// TIA Portal project "Delta_Praktika_P&P" (V17) (continued)
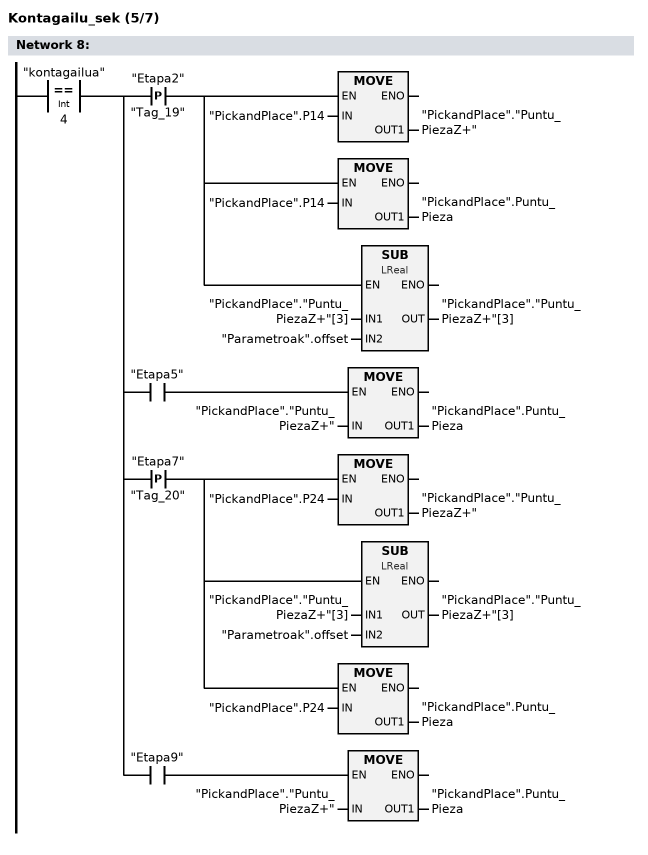
   RUNG wire#powerrail
      { S7_Templates := "SrcType := Int" } EQ_Contact(in1 := "kontagailua", in2 := 4)
      wire#w1
      P_Contact(operand := "Etapa2", bit := "Tag_19")
      wire#w2
      Move(in := "PickandPlace".P14, out1 => "PickandPlace"."Puntu_PiezaZ+")
   END_RUNG
   RUNG wire#w2
      Move(in := "PickandPlace".P14, out1 => "PickandPlace".Puntu_Pieza)
   END_RUNG
   RUNG wire#w2
      { S7_Templates := "SrcType := LReal" } Sub(in1 := "PickandPlace"."Puntu_PiezaZ+"[3], in2 := "Parametroak".offset, out => "PickandPlace"."Puntu_PiezaZ+"[3])
   END_RUNG
   RUNG wire#w1
      Contact( "Etapa5" )
      Move(in := "PickandPlace"."Puntu_PiezaZ+", out1 => "PickandPlace".Puntu_Pieza)
   END_RUNG
   RUNG wire#w1
      P_Contact(operand := "Etapa7", bit := "Tag_20")
      wire#w3
      Move(in := "PickandPlace".P24, out1 => "PickandPlace"."Puntu_PiezaZ+")
   END_RUNG
   RUNG wire#w3
      { S7_Templates := "SrcType := LReal" } Sub(in1 := "PickandPlace"."Puntu_PiezaZ+"[3], in2 := "Parametroak".offset, out => "PickandPlace"."Puntu_PiezaZ+"[3])
   END_RUNG
   RUNG wire#w3
      Move(in := "PickandPlace".P24, out1 => "PickandPlace".Puntu_Pieza)
   END_RUNG
   RUNG wire#w1
      Contact( "Etapa9" )
      Move(in := "PickandPlace"."Puntu_PiezaZ+", out1 => "PickandPlace".Puntu_Pieza)
   END_RUNG
   // the same network as SCL:
   #_w1 := "kontagailua" = 4;
   #_w2 := #_w1 AND "Etapa2" AND NOT "Tag_19";   // rising edge of "Etapa2"
   "Tag_19" := "Etapa2";
   IF #_w2 THEN
       "PickandPlace"."Puntu_PiezaZ+" := "PickandPlace".P14;
       "PickandPlace".Puntu_Pieza := "PickandPlace".P14;
       "PickandPlace"."Puntu_PiezaZ+"[3] := "PickandPlace"."Puntu_PiezaZ+"[3] - "Parametroak".offset;
   END_IF;
   IF #_w1 AND "Etapa5" THEN "PickandPlace".Puntu_Pieza := "PickandPlace"."Puntu_PiezaZ+"; END_IF;
   #_w3 := #_w1 AND "Etapa7" AND NOT "Tag_20";   // rising edge of "Etapa7"
   "Tag_20" := "Etapa7";
   IF #_w3 THEN
       "PickandPlace"."Puntu_PiezaZ+" := "PickandPlace".P24;
       "PickandPlace"."Puntu_PiezaZ+"[3] := "PickandPlace"."Puntu_PiezaZ+"[3] - "Parametroak".offset;
       "PickandPlace".Puntu_Pieza := "PickandPlace".P24;
   END_IF;
   IF #_w1 AND "Etapa9" THEN "PickandPlace".Puntu_Pieza := "PickandPlace"."Puntu_PiezaZ+"; END_IF;
END_REGION

REGION Network 9
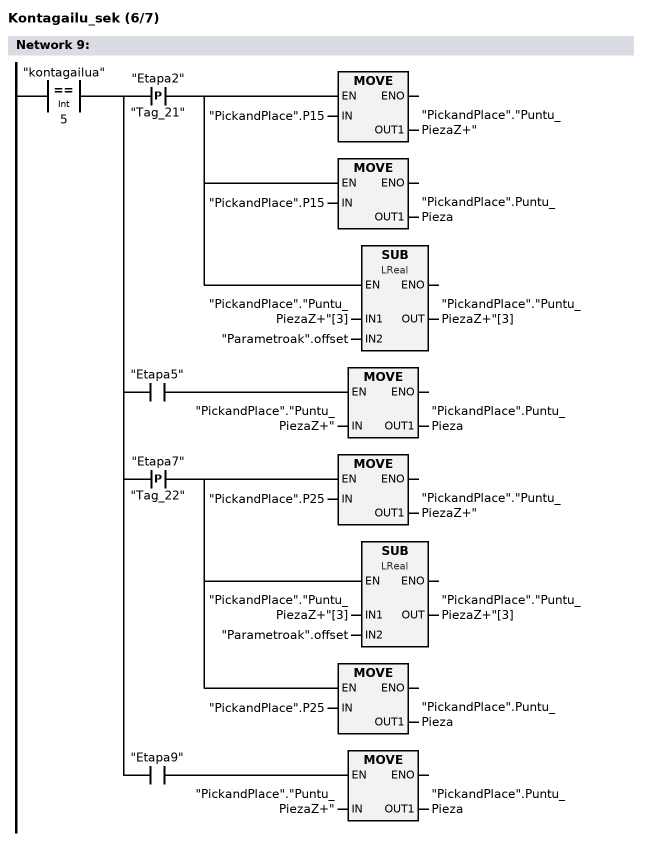
   RUNG wire#powerrail
      { S7_Templates := "SrcType := Int" } EQ_Contact(in1 := "kontagailua", in2 := 5)
      wire#w1
      P_Contact(operand := "Etapa2", bit := "Tag_21")
      wire#w2
      Move(in := "PickandPlace".P15, out1 => "PickandPlace"."Puntu_PiezaZ+")
   END_RUNG
   RUNG wire#w2
      Move(in := "PickandPlace".P15, out1 => "PickandPlace".Puntu_Pieza)
   END_RUNG
   RUNG wire#w2
      { S7_Templates := "SrcType := LReal" } Sub(in1 := "PickandPlace"."Puntu_PiezaZ+"[3], in2 := "Parametroak".offset, out => "PickandPlace"."Puntu_PiezaZ+"[3])
   END_RUNG
   RUNG wire#w1
      Contact( "Etapa5" )
      Move(in := "PickandPlace"."Puntu_PiezaZ+", out1 => "PickandPlace".Puntu_Pieza)
   END_RUNG
   RUNG wire#w1
      P_Contact(operand := "Etapa7", bit := "Tag_22")
      wire#w3
      Move(in := "PickandPlace".P25, out1 => "PickandPlace"."Puntu_PiezaZ+")
   END_RUNG
   RUNG wire#w3
      { S7_Templates := "SrcType := LReal" } Sub(in1 := "PickandPlace"."Puntu_PiezaZ+"[3], in2 := "Parametroak".offset, out => "PickandPlace"."Puntu_PiezaZ+"[3])
   END_RUNG
   RUNG wire#w3
      Move(in := "PickandPlace".P25, out1 => "PickandPlace".Puntu_Pieza)
   END_RUNG
   RUNG wire#w1
      Contact( "Etapa9" )
      Move(in := "PickandPlace"."Puntu_PiezaZ+", out1 => "PickandPlace".Puntu_Pieza)
   END_RUNG
   // the same network as SCL:
   #_w1 := "kontagailua" = 5;
   #_w2 := #_w1 AND "Etapa2" AND NOT "Tag_21";   // rising edge of "Etapa2"
   "Tag_21" := "Etapa2";
   IF #_w2 THEN
       "PickandPlace"."Puntu_PiezaZ+" := "PickandPlace".P15;
       "PickandPlace".Puntu_Pieza := "PickandPlace".P15;
       "PickandPlace"."Puntu_PiezaZ+"[3] := "PickandPlace"."Puntu_PiezaZ+"[3] - "Parametroak".offset;
   END_IF;
   IF #_w1 AND "Etapa5" THEN "PickandPlace".Puntu_Pieza := "PickandPlace"."Puntu_PiezaZ+"; END_IF;
   #_w3 := #_w1 AND "Etapa7" AND NOT "Tag_22";   // rising edge of "Etapa7"
   "Tag_22" := "Etapa7";
   IF #_w3 THEN
       "PickandPlace"."Puntu_PiezaZ+" := "PickandPlace".P25;
       "PickandPlace"."Puntu_PiezaZ+"[3] := "PickandPlace"."Puntu_PiezaZ+"[3] - "Parametroak".offset;
       "PickandPlace".Puntu_Pieza := "PickandPlace".P25;
   END_IF;
   IF #_w1 AND "Etapa9" THEN "PickandPlace".Puntu_Pieza := "PickandPlace"."Puntu_PiezaZ+"; END_IF;
END_REGION

REGION Network 10
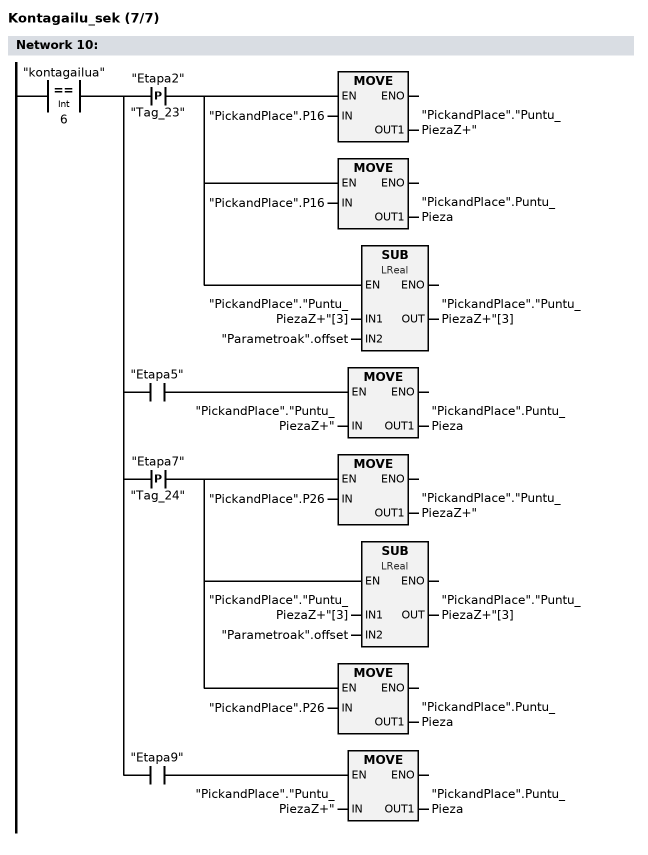
   RUNG wire#powerrail
      { S7_Templates := "SrcType := Int" } EQ_Contact(in1 := "kontagailua", in2 := 6)
      wire#w1
      P_Contact(operand := "Etapa2", bit := "Tag_23")
      wire#w2
      Move(in := "PickandPlace".P16, out1 => "PickandPlace"."Puntu_PiezaZ+")
   END_RUNG
   RUNG wire#w2
      Move(in := "PickandPlace".P16, out1 => "PickandPlace".Puntu_Pieza)
   END_RUNG
   RUNG wire#w2
      { S7_Templates := "SrcType := LReal" } Sub(in1 := "PickandPlace"."Puntu_PiezaZ+"[3], in2 := "Parametroak".offset, out => "PickandPlace"."Puntu_PiezaZ+"[3])
   END_RUNG
   RUNG wire#w1
      Contact( "Etapa5" )
      Move(in := "PickandPlace"."Puntu_PiezaZ+", out1 => "PickandPlace".Puntu_Pieza)
   END_RUNG
   RUNG wire#w1
      P_Contact(operand := "Etapa7", bit := "Tag_24")
      wire#w3
      Move(in := "PickandPlace".P26, out1 => "PickandPlace"."Puntu_PiezaZ+")
   END_RUNG
   RUNG wire#w3
      { S7_Templates := "SrcType := LReal" } Sub(in1 := "PickandPlace"."Puntu_PiezaZ+"[3], in2 := "Parametroak".offset, out => "PickandPlace"."Puntu_PiezaZ+"[3])
   END_RUNG
   RUNG wire#w3
      Move(in := "PickandPlace".P26, out1 => "PickandPlace".Puntu_Pieza)
   END_RUNG
   RUNG wire#w1
      Contact( "Etapa9" )
      Move(in := "PickandPlace"."Puntu_PiezaZ+", out1 => "PickandPlace".Puntu_Pieza)
   END_RUNG
   // the same network as SCL:
   #_w1 := "kontagailua" = 6;
   #_w2 := #_w1 AND "Etapa2" AND NOT "Tag_23";   // rising edge of "Etapa2"
   "Tag_23" := "Etapa2";
   IF #_w2 THEN
       "PickandPlace"."Puntu_PiezaZ+" := "PickandPlace".P16;
       "PickandPlace".Puntu_Pieza := "PickandPlace".P16;
       "PickandPlace"."Puntu_PiezaZ+"[3] := "PickandPlace"."Puntu_PiezaZ+"[3] - "Parametroak".offset;
   END_IF;
   IF #_w1 AND "Etapa5" THEN "PickandPlace".Puntu_Pieza := "PickandPlace"."Puntu_PiezaZ+"; END_IF;
   #_w3 := #_w1 AND "Etapa7" AND NOT "Tag_24";   // rising edge of "Etapa7"
   "Tag_24" := "Etapa7";
   IF #_w3 THEN
       "PickandPlace"."Puntu_PiezaZ+" := "PickandPlace".P26;
       "PickandPlace"."Puntu_PiezaZ+"[3] := "PickandPlace"."Puntu_PiezaZ+"[3] - "Parametroak".offset;
       "PickandPlace".Puntu_Pieza := "PickandPlace".P26;
   END_IF;
   IF #_w1 AND "Etapa9" THEN "PickandPlace".Puntu_Pieza := "PickandPlace"."Puntu_PiezaZ+"; END_IF;
END_REGION
END_FUNCTION

ORGANIZATION_BLOCK "Main"   // OB1, LAD, ProgramCycle
TITLE = "Main Program Sweep (Cycle)"
{ S7_Optimized_Access := 'TRUE' }
VERSION : 0.1
   VAR_INPUT
      Initial_Call : Bool;   // Initial call of this OB
      Remanence : Bool;   // =True, if remanent data are available
   END_VAR
BEGIN

REGION Network 1
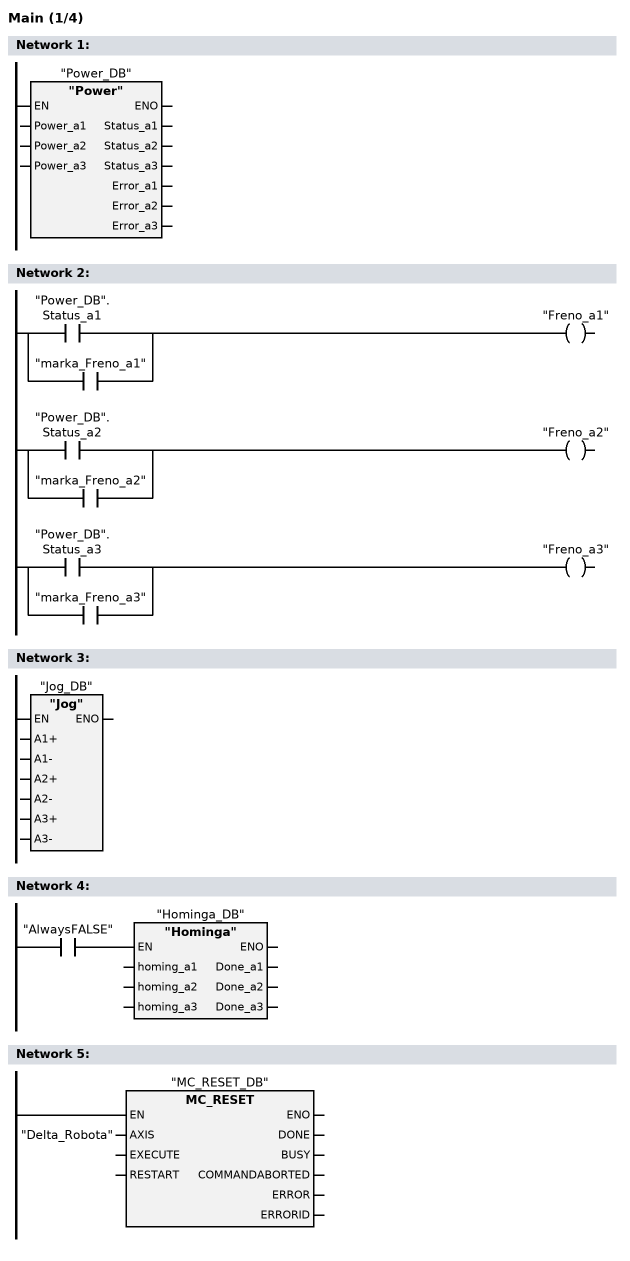
   RUNG wire#powerrail
      "Power_DB"(Power_a1 :=, Power_a2 :=, Power_a3 :=, Status_a1 =>, Status_a2 =>, Status_a3 =>, Error_a1 =>, Error_a2 =>, Error_a3 =>)
   END_RUNG
   // the same network as SCL:
   "Power_DB"();   // "Power"
END_REGION

REGION Network 2
   RUNG wire#powerrail
      Contact( "Power_DB".Status_a1 )
      wire#w1
      Coil( "Freno_a1" )
   END_RUNG
   RUNG wire#powerrail
      Contact( "marka_Freno_a1" )
   END_RUNG wire#w1
   RUNG wire#powerrail
      Contact( "Power_DB".Status_a2 )
      wire#w2
      Coil( "Freno_a2" )
   END_RUNG
   RUNG wire#powerrail
      Contact( "marka_Freno_a2" )
   END_RUNG wire#w2
   RUNG wire#powerrail
      Contact( "Power_DB".Status_a3 )
      wire#w3
      Coil( "Freno_a3" )
   END_RUNG
   RUNG wire#powerrail
      Contact( "marka_Freno_a3" )
   END_RUNG wire#w3
   // the same network as SCL:
   "Freno_a1" := "Power_DB".Status_a1 OR "marka_Freno_a1";
   "Freno_a2" := "Power_DB".Status_a2 OR "marka_Freno_a2";
   "Freno_a3" := "Power_DB".Status_a3 OR "marka_Freno_a3";
END_REGION

REGION Network 3
   RUNG wire#powerrail
      "Jog_DB"("A1+" :=, "A1-" :=, "A2+" :=, "A2-" :=, "A3+" :=, "A3-" :=)
   END_RUNG
   // the same network as SCL:
   "Jog_DB"();   // "Jog"
END_REGION

REGION Network 4
   RUNG wire#powerrail
      Contact( "AlwaysFALSE" )
      "Hominga_DB"(homing_a1 :=, homing_a2 :=, homing_a3 :=, Done_a1 =>, Done_a2 =>, Done_a3 =>)
   END_RUNG
   // the same network as SCL:
   IF "AlwaysFALSE" THEN
       "Hominga_DB"();   // "Hominga"
   END_IF;
END_REGION

REGION Network 5
   "MC_RESET_DB"(Axis := "Delta_Robota");   // MC_RESET
END_REGION

REGION Network 6
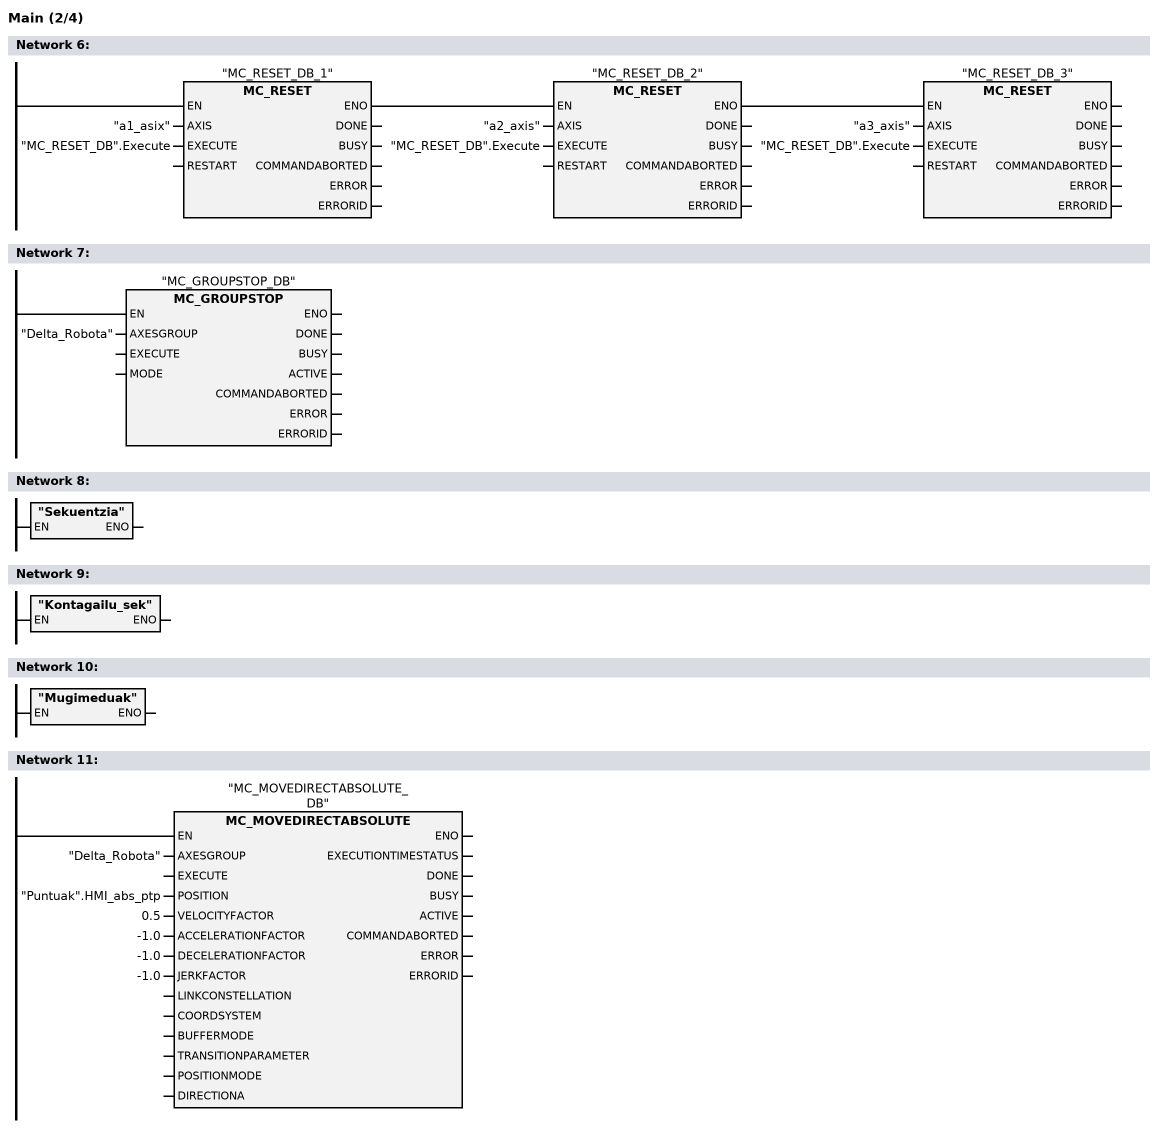
   // ENO of a box is taken as its EN; it also drops when the box reports an error
   "MC_RESET_DB_1"(Axis := "a1_asix", Execute := "MC_RESET_DB".Execute);   // MC_RESET
   "MC_RESET_DB_2"(Axis := "a2_axis", Execute := "MC_RESET_DB".Execute);   // MC_RESET
   "MC_RESET_DB_3"(Axis := "a3_axis", Execute := "MC_RESET_DB".Execute);   // MC_RESET
END_REGION

REGION Network 7
   "MC_GROUPSTOP_DB"(AxesGroup := "Delta_Robota");   // MC_GROUPSTOP
END_REGION

REGION Network 8
   RUNG wire#powerrail
      "Sekuentzia"()
   END_RUNG
   // the same network as SCL:
   "Sekuentzia"();
END_REGION

REGION Network 9
   RUNG wire#powerrail
      "Kontagailu_sek"()
   END_RUNG
   // the same network as SCL:
   "Kontagailu_sek"();
END_REGION

REGION Network 10
   RUNG wire#powerrail
      "Mugimeduak"()
   END_RUNG
   // the same network as SCL:
   "Mugimeduak"();
END_REGION

REGION Network 11
   "MC_MOVEDIRECTABSOLUTE_DB"(AxesGroup := "Delta_Robota",   // MC_MOVEDIRECTABSOLUTE
                           Position := "Puntuak".HMI_abs_ptp,
                           VelocityFactor := 0.5,
                           AccelerationFactor := -1.0,
                           DecelerationFactor := -1.0,
                           JerkFactor := -1.0);
END_REGION

REGION Network 12
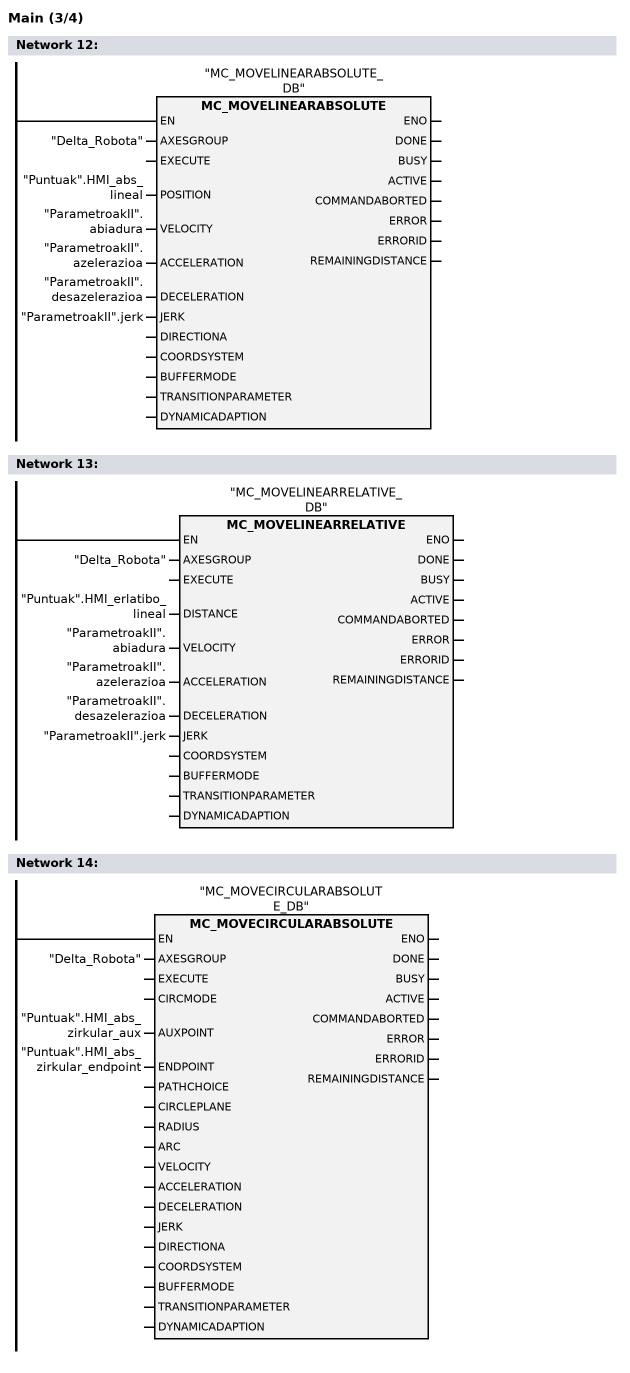
   "MC_MOVELINEARABSOLUTE_DB"(AxesGroup := "Delta_Robota",   // MC_MOVELINEARABSOLUTE
                           Position := "Puntuak".HMI_abs_lineal,
                           Velocity := "ParametroakII".abiadura,
                           Acceleration := "ParametroakII".azelerazioa,
                           Deceleration := "ParametroakII".desazelerazioa,
                           Jerk := "ParametroakII".jerk);
END_REGION

REGION Network 13
   "MC_MOVELINEARRELATIVE_DB"(AxesGroup := "Delta_Robota",   // MC_MOVELINEARRELATIVE
                           Distance := "Puntuak".HMI_erlatibo_lineal,
                           Velocity := "ParametroakII".abiadura,
                           Acceleration := "ParametroakII".azelerazioa,
                           Deceleration := "ParametroakII".desazelerazioa,
                           Jerk := "ParametroakII".jerk);
END_REGION

REGION Network 14
   "MC_MOVECIRCULARABSOLUTE_DB"(AxesGroup := "Delta_Robota",   // MC_MOVECIRCULARABSOLUTE
                           AuxPoint := "Puntuak".HMI_abs_zirkular_aux,
                           EndPoint := "Puntuak".HMI_abs_zirkular_endpoint);
END_REGION

REGION Network 15
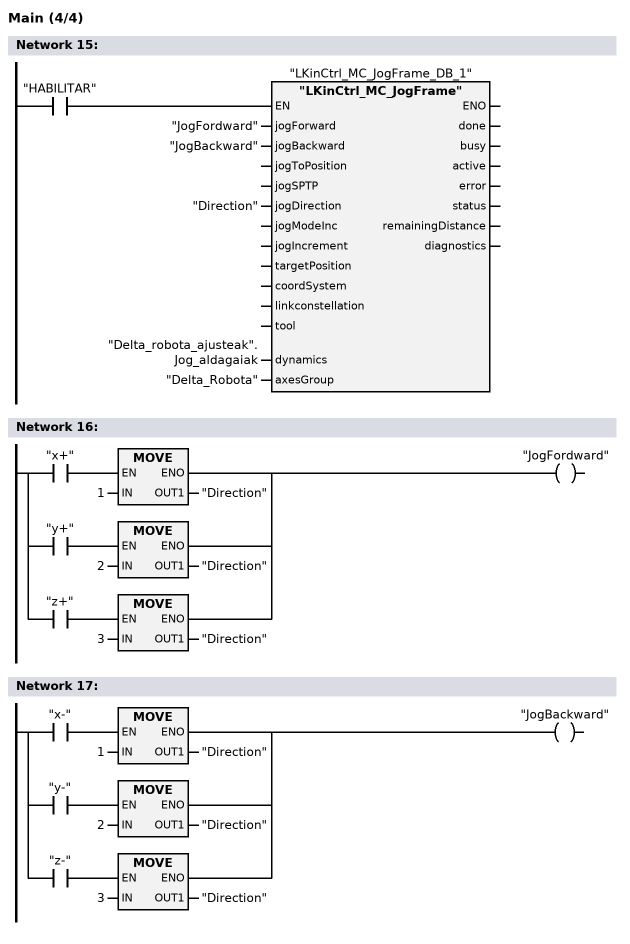
   RUNG wire#powerrail
      Contact( "HABILITAR" )
      "LKinCtrl_MC_JogFrame_DB_1"(jogForward := "JogFordward", jogBackward := "JogBackward", jogToPosition :=, jogSPTP :=, jogDirection := "Direction", jogModeInc :=, jogIncrement :=, targetPosition :=, coordSystem :=, linkconstellation :=, tool :=, dynamics := "Delta_robota_ajusteak".Jog_aldagaiak, axesGroup := "Delta_Robota", done =>, busy =>, active =>, error =>, status =>, remainingDistance =>, diagnostics =>)
   END_RUNG
   // the same network as SCL:
   IF "HABILITAR" THEN
       "LKinCtrl_MC_JogFrame_DB_1"(jogForward := "JogFordward",   // "LKinCtrl_MC_JogFrame"
                               jogBackward := "JogBackward",
                               jogDirection := "Direction",
                               dynamics := "Delta_robota_ajusteak".Jog_aldagaiak,
                               axesGroup := "Delta_Robota");
   END_IF;
END_REGION

REGION Network 16
   RUNG wire#powerrail
      Contact( "x+" )
      Move(in := 1, out1 => "Direction")
      wire#w1
      Coil( "JogFordward" )
   END_RUNG
   RUNG wire#powerrail
      Contact( "y+" )
      Move(in := 2, out1 => "Direction")
   END_RUNG wire#w1
   RUNG wire#powerrail
      Contact( "z+" )
      Move(in := 3, out1 => "Direction")
   END_RUNG wire#w1
   // the same network as SCL:
   IF "x+" THEN "Direction" := 1; END_IF;
   IF "y+" THEN "Direction" := 2; END_IF;
   IF "z+" THEN "Direction" := 3; END_IF;
   "JogFordward" := "x+" OR "y+" OR "z+";
END_REGION

REGION Network 17
   RUNG wire#powerrail
      Contact( "x-" )
      Move(in := 1, out1 => "Direction")
      wire#w1
      Coil( "JogBackward" )
   END_RUNG
   RUNG wire#powerrail
      Contact( "y-" )
      Move(in := 2, out1 => "Direction")
   END_RUNG wire#w1
   RUNG wire#powerrail
      Contact( "z-" )
      Move(in := 3, out1 => "Direction")
   END_RUNG wire#w1
   // the same network as SCL:
   IF "x-" THEN "Direction" := 1; END_IF;
   IF "y-" THEN "Direction" := 2; END_IF;
   IF "z-" THEN "Direction" := 3; END_IF;
   "JogBackward" := "x-" OR "y-" OR "z-";
END_REGION
END_ORGANIZATION_BLOCK

ORGANIZATION_BLOCK "Startup"   // OB100, LAD, Startup
TITLE = "Complete Restart"
{ S7_Optimized_Access := 'TRUE' }
VERSION : 0.1
   VAR_INPUT
      LostRetentive : Bool;   // True if retentive data are lost
      LostRTC : Bool;   // True if date and time are lost
   END_VAR
BEGIN

REGION Network 1
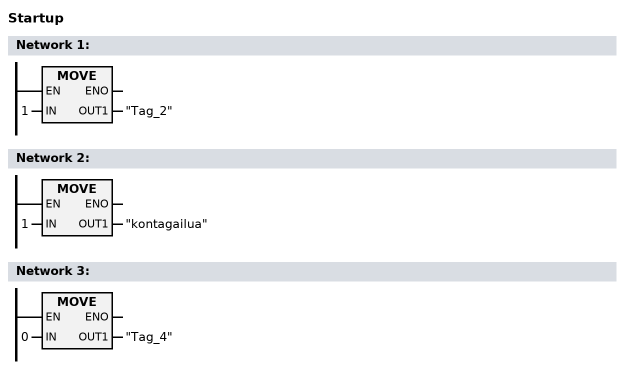
   RUNG wire#powerrail
      Move(in := 1, out1 => "Tag_2")
   END_RUNG
   // the same network as SCL:
   "Tag_2" := 1;
END_REGION

REGION Network 2
   RUNG wire#powerrail
      Move(in := 1, out1 => "kontagailua")
   END_RUNG
   // the same network as SCL:
   "kontagailua" := 1;
END_REGION

REGION Network 3
   RUNG wire#powerrail
      Move(in := 0, out1 => "Tag_4")
   END_RUNG
   // the same network as SCL:
   "Tag_4" := 0;
END_REGION
END_ORGANIZATION_BLOCK

(* ===== HMI "HMI_RT_1" =====
system functions are stored by id; their names below are inferred from use
connection "HMI_Conexión_2": ETHERNET, SMART_S7_1500_OMS

HMI tags "Tabla de variables estándar"
   "Delta_Robota_TcpInWcs_x_Position" : LReal = PLC Delta_Robota.TcpInWcs.x.Position, 1 s
   "Power_DB_Power_a1" : Bool = PLC Power_DB.Power_a1, 1 s
   "Jog_DB_A1+" : Bool = PLC Jog_DB.A1+, 1 s
   "a1_asix_ActualPosition" : LReal = PLC a1_asix.ActualPosition, 1 s
   "Power_DB_Power_a2" : Bool = PLC Power_DB.Power_a2, 1 s
   "Power_DB_Power_a3" : Bool = PLC Power_DB.Power_a3, 1 s
   "Tag_2" : Bool = PLC marka_Freno_a1 AT %M30.1, 1 s
   "Tag_3" : Bool = PLC marka_Freno_a2 AT %M30.2, 1 s
   "Tag_6" : Bool = PLC marka_Freno_a3 AT %M30.0, 1 s
   "Jog_DB_A1-" : Bool = PLC Jog_DB.A1-, 1 s
   "Jog_DB_A2+" : Bool = PLC Jog_DB.A2+, 1 s
   "Jog_DB_A2-" : Bool = PLC Jog_DB.A2-, 1 s
   "Jog_DB_A3+" : Bool = PLC Jog_DB.A3+, 1 s
   "Jog_DB_A3-" : Bool = PLC Jog_DB.A3-, 1 s
   "Tag_1" : Bool = PLC Freno_a1 AT %Q30.1, 1 s
   "Tag_4" : Bool = PLC Freno_a2 AT %Q30.2, 1 s
   "a3_axis_ActualPosition" : LReal = PLC a3_axis.ActualPosition, 1 s
   "Tag_5" : Bool = PLC Freno_a3 AT %Q30.0, 1 s
   "Delta_Robota_TcpInWcs_y_Position" : LReal = PLC Delta_Robota.TcpInWcs.y.Position, 1 s
   "Delta_Robota_TcpInWcs_z_Position" : LReal = PLC Delta_Robota.TcpInWcs.z.Position, 1 s
   "a2_axis_ActualPosition" : LReal = PLC a2_axis.ActualPosition, 1 s
   "MC_GROUPSTOP_DB_Execute" : Bool = PLC MC_GROUPSTOP_DB.Execute, 1 s
   "MC_RESET_DB_Execute" : Bool = PLC MC_RESET_DB.Execute, 1 s
   "Puntuak_HMI_erlatibo_lineal{1}" : LReal = PLC Puntuak.HMI_erlatibo_lineal[1], 1 s
   "Puntuak_HMI_erlatibo_lineal{2}" : LReal = PLC Puntuak.HMI_erlatibo_lineal[2], 1 s
   "Puntuak_HMI_erlatibo_lineal{3}" : LReal = PLC Puntuak.HMI_erlatibo_lineal[3], 1 s
   "Puntuak_HMI_abs_lineal{1}" : LReal = PLC Puntuak.HMI_abs_lineal[1], 1 s
   "Puntuak_HMI_abs_lineal{2}" : LReal = PLC Puntuak.HMI_abs_lineal[2], 1 s
   "Puntuak_HMI_abs_lineal{3}" : LReal = PLC Puntuak.HMI_abs_lineal[3], 1 s
   "Puntuak_HMI_abs_ptp{1}" : LReal = PLC Puntuak.HMI_abs_ptp[1], 1 s
   "Puntuak_HMI_abs_ptp{2}" : LReal = PLC Puntuak.HMI_abs_ptp[2], 1 s
   "Puntuak_HMI_abs_ptp{3}" : LReal = PLC Puntuak.HMI_abs_ptp[3], 1 s
   "MC_MOVELINEARABSOLUTE_DB_Execute" : Bool = PLC MC_MOVELINEARABSOLUTE_DB.Execute, 1 s
   "MC_MOVEDIRECTABSOLUTE_DB_Execute" : Bool = PLC MC_MOVEDIRECTABSOLUTE_DB.Execute, 1 s
   "MC_MOVELINEARRELATIVE_DB_Execute" : Bool = PLC MC_MOVELINEARRELATIVE_DB.Execute, 1 s
   "Puntuak_HMI_abs_zirkular_aux{1}" : LReal = PLC Puntuak.HMI_abs_zirkular_aux[1], 1 s
   "Puntuak_HMI_abs_zirkular_aux{2}" : LReal = PLC Puntuak.HMI_abs_zirkular_aux[2], 1 s
   "Puntuak_HMI_abs_zirkular_aux{3}" : LReal = PLC Puntuak.HMI_abs_zirkular_aux[3], 1 s
   "Puntuak_HMI_abs_zirkular_endpoint{1}" : LReal = PLC Puntuak.HMI_abs_zirkular_endpoint[1], 1 s
   "Puntuak_HMI_abs_zirkular_endpoint{2}" : LReal = PLC Puntuak.HMI_abs_zirkular_endpoint[2], 1 s
   "Puntuak_HMI_abs_zirkular_endpoint{3}" : LReal = PLC Puntuak.HMI_abs_zirkular_endpoint[3], 1 s
   "MC_MOVECIRCULARABSOLUTE_DB_Execute" : Bool = PLC MC_MOVECIRCULARABSOLUTE_DB.Execute, 1 s
   "HABILITAR" : Bool = PLC HABILITAR AT %M150.2, 1 s
   "x+" : Bool = PLC "x+" AT %M152.0, 1 s
   "x-" : Bool = PLC "x-" AT %M152.1, 1 s
   "y+" : Bool = PLC "y+" AT %M152.2, 1 s
   "y-" : Bool = PLC "y-" AT %M152.3, 1 s
   "z+" : Bool = PLC "z+" AT %M152.4, 1 s
   "z-" : Bool = PLC "z-" AT %M152.5, 1 s
   "HMI_start" : Bool = PLC HMI_start AT %M10.0, 1 s

screen "Imagen_1" 1280x800
   Button "Botón_1" at 38,159 size 96x32; TextOff 'A1+'
      on Press: function_b14e0dd5("Jog_DB_A1+", 0)
   Button "Botón_2" at 175,159 size 96x32; TextOff 'A1-'
      on Press: function_b14e0dd5("Jog_DB_A1-", 0)
   Button "Botón_3" at 40,207 size 96x32; TextOff 'A2+'
      on Press: function_b14e0dd5("Jog_DB_A2+", 0)
   Button "Botón_4" at 175,207 size 96x32; TextOff 'A2-'
      on Press: function_b14e0dd5("Jog_DB_A2-", 0)
   Button "Botón_5" at 40,255 size 96x32; TextOff 'A3+'
      on Press: function_b14e0dd5("Jog_DB_A3+", 0)
   Button "Botón_6" at 175,255 size 96x32; TextOff 'A3-'
      on Press: function_b14e0dd5("Jog_DB_A3-", 0)
   Button "Botón_10" at 926,70 size 96x32; TextOff 'Stop'
      on Press: function_b14e0dd5("MC_GROUPSTOP_DB_Execute", 0)
   Button "Botón_11" at 1061,70 size 96x32; TextOff 'Reset'
      on Press: function_b14e0dd5("MC_RESET_DB_Execute", 0)
   TextField "Campo de texto_1" at 68,12 size 306x23; Text 'OBJETO TEKNOLOGIKOA BANAKA'
   TextField "Campo de texto_2" at 850,14 size 146x23; Text 'DELTA ROBOTA'
   Circle "Círculo_1" at 415,164 size 19x19
      Appearance <- "Tag_1"
   Circle "Círculo_2" at 415,212 size 19x19
      Appearance <- "Tag_4"
   Circle "Círculo_3" at 415,260 size 19x19
      Appearance <- "Tag_5"
   TextField "Campo de texto_3" at 144,116 size 330x23; Text 'Frenoa desaktibatuta badago berde'
   IOField "Campo ES_1" at 921,418 size 80x30; FormatPattern s999.99
      ProcessValue <- "Puntuak_HMI_abs_lineal{1}"
   IOField "Campo ES_2" at 920,452 size 81x30; FormatPattern s999.99
      ProcessValue <- "Puntuak_HMI_abs_lineal{2}"
   IOField "Campo ES_3" at 920,486 size 81x33; FormatPattern s999.99
      ProcessValue <- "Puntuak_HMI_abs_lineal{3}"
   Button "Botón_15" at 1048,454 size 96x32; TextOff 'GO!'
      on Press: function_b14e0dd5("MC_MOVELINEARABSOLUTE_DB_Execute", 0)
   TextField "Campo de texto_4" at 928,382 size 270x23; Text 'Mugimendu absoluto linearra'
   TextField "Campo de texto_5" at 1001,418 size 47x23; Text 'X'
   TextField "Campo de texto_6" at 1001,455 size 47x23; Text 'Y'
   TextField "Campo de texto_7" at 1001,492 size 47x23; Text 'Z'
   IOField "Campo ES_4" at 959,607 size 73x30; FormatPattern 99999
   IOField "Campo ES_5" at 959,641 size 73x30; FormatPattern 99999
   IOField "Campo ES_6" at 959,675 size 73x30; FormatPattern 99999
   Button "Botón_16" at 1017,715 size 96x32; TextOff 'GO!'
   TextField "Campo de texto_8" at 959,545 size 288x23; Text 'Mugimendu absoluto zirkularra'
   TextField "Campo de texto_9" at 1032,607 size 47x23; Text 'X'
   TextField "Campo de texto_10" at 1032,644 size 47x23; Text 'Y'
   TextField "Campo de texto_11" at 1032,681 size 47x23; Text 'Z'
   IOField "Campo ES_7" at 1083,608 size 73x30; FormatPattern 99999
   IOField "Campo ES_8" at 1083,642 size 73x30; FormatPattern 99999
   IOField "Campo ES_9" at 1083,676 size 73x30; FormatPattern 99999
   TextField "Campo de texto_12" at 1159,608 size 47x23; Text 'X'
   TextField "Campo de texto_13" at 1159,645 size 47x23; Text 'Y'
   TextField "Campo de texto_14" at 1159,682 size 47x23; Text 'Z'
   TextField "Campo de texto_15" at 928,575 size 135x23; Text 'Nundik pasatu'
   TextField "Campo de texto_16" at 1079,575 size 142x23; Text 'Azken posizioa'
   IOField "Campo ES_13" at 954,607 size 78x31; FormatPattern s999.99
      ProcessValue <- "Puntuak_HMI_abs_zirkular_aux{1}"
   IOField "Campo ES_14" at 954,641 size 78x30; FormatPattern s999.99
      ProcessValue <- "Puntuak_HMI_abs_zirkular_aux{2}"
   IOField "Campo ES_15" at 952,675 size 80x30; FormatPattern s999.99
      ProcessValue <- "Puntuak_HMI_abs_zirkular_aux{3}"
   Button "Botón_18" at 1017,715 size 96x32; TextOff 'GO!'
      on Press: function_b14e0dd5("MC_MOVECIRCULARABSOLUTE_DB_Execute", 0)
   TextField "Campo de texto_21" at 959,545 size 288x23; Text 'Mugimendu absoluto zirkularra'
   TextField "Campo de texto_22" at 1032,607 size 47x23; Text 'X'
   TextField "Campo de texto_23" at 1032,644 size 47x23; Text 'Y'
   TextField "Campo de texto_24" at 1032,681 size 47x23; Text 'Z'
   IOField "Campo ES_16" at 1077,608 size 79x30; FormatPattern s999.99
      ProcessValue <- "Puntuak_HMI_abs_zirkular_endpoint{1}"
   IOField "Campo ES_17" at 1078,642 size 78x30; FormatPattern s999.99
      ProcessValue <- "Puntuak_HMI_abs_zirkular_endpoint{2}"
   IOField "Campo ES_18" at 1078,676 size 78x30; FormatPattern s999.99
      ProcessValue <- "Puntuak_HMI_abs_zirkular_endpoint{3}"
   TextField "Campo de texto_25" at 1159,608 size 47x23; Text 'X'
   TextField "Campo de texto_26" at 1159,645 size 47x23; Text 'Y'
   TextField "Campo de texto_27" at 1159,682 size 47x23; Text 'Z'
   TextField "Campo de texto_28" at 928,575 size 135x23; Text 'Nundik pasatu'
   TextField "Campo de texto_29" at 1079,575 size 142x23; Text 'Azken posizioa'
   IOField "Campo ES_10" at 40,390 size 96x32; FormatPattern s99.999
      ProcessValue <- "a1_asix_ActualPosition"
   IOField "Campo ES_11" at 166,388 size 96x32; FormatPattern s99.999
      ProcessValue <- "a2_axis_ActualPosition"
   IOField "Campo ES_12" at 308,388 size 96x32; FormatPattern s99.999
      ProcessValue <- "a3_axis_ActualPosition"
   TextField "Campo de texto_17" at 68,352 size 46x25; Text 'A1'
   TextField "Campo de texto_18" at 198,352 size 46x25; Text 'A2'
   TextField "Campo de texto_19" at 328,352 size 46x25; Text 'A3'
   IOField "Campo ES_19" at 549,418 size 86x33; FormatPattern s999.99
      ProcessValue <- "Puntuak_HMI_erlatibo_lineal{1}"
   IOField "Campo ES_20" at 550,452 size 85x31; FormatPattern s999.99
      ProcessValue <- "Puntuak_HMI_erlatibo_lineal{2}"
   IOField "Campo ES_21" at 550,486 size 85x30; FormatPattern s999.99
      ProcessValue <- "Puntuak_HMI_erlatibo_lineal{3}"
   Button "Botón_17" at 682,454 size 96x32; TextOff 'GO!'
      on Press: function_b14e0dd5("MC_MOVELINEARRELATIVE_DB_Execute", 0)
   TextField "Campo de texto_20" at 562,382 size 264x23; Text 'Mugimendu erlatibo linearra'
   TextField "Campo de texto_30" at 635,418 size 47x23; Text 'X'
   TextField "Campo de texto_31" at 635,455 size 47x23; Text 'Y'
   TextField "Campo de texto_32" at 635,492 size 47x23; Text 'Z'
   IOField "Campo ES_25" at 594,613 size 73x30; FormatPattern 99999
   IOField "Campo ES_26" at 594,647 size 73x30; FormatPattern 99999
   IOField "Campo ES_27" at 594,681 size 73x30; FormatPattern 99999
   TextField "Campo de texto_37" at 682,618 size 47x23; Text 'X'
   TextField "Campo de texto_38" at 682,655 size 47x23; Text 'Y'
   TextField "Campo de texto_39" at 682,692 size 47x23; Text 'Z'
   Button "Botón_20" at 713,649 size 96x32; TextOff 'GO!'
      on Press: function_b14e0dd5("MC_MOVEDIRECTABSOLUTE_DB_Execute", 0)
   IOField "Campo ES_31" at 585,613 size 82x31; FormatPattern s999.99
      ProcessValue <- "Puntuak_HMI_abs_ptp{1}"
   IOField "Campo ES_32" at 584,647 size 83x31; FormatPattern s999.99
      ProcessValue <- "Puntuak_HMI_abs_ptp{2}"
   IOField "Campo ES_33" at 584,681 size 83x29; FormatPattern s999.99
      ProcessValue <- "Puntuak_HMI_abs_ptp{3}"
   TextField "Campo de texto_46" at 682,618 size 47x23; Text 'X'
   TextField "Campo de texto_47" at 682,655 size 47x23; Text 'Y'
   TextField "Campo de texto_48" at 682,692 size 47x23; Text 'Z'
   TextField "Campo de texto_42" at 581,326 size 254x25; Text 'MUGIMENDU ERLATIBOAK'
   TextField "Campo de texto_51" at 603,540 size 261x25; Text 'MUGIMENDU ABSOLUTOAK'
   IOField "Campo ES_34" at 520,119 size 108x32; FormatPattern s999.999
      ProcessValue <- "Delta_Robota_TcpInWcs_x_Position"
   IOField "Campo ES_35" at 520,179 size 108x33; FormatPattern s999.999
      ProcessValue <- "Delta_Robota_TcpInWcs_y_Position"
   IOField "Campo ES_36" at 521,239 size 107x35; FormatPattern s999.999
      ProcessValue <- "Delta_Robota_TcpInWcs_z_Position"
   TextField "Campo de texto_52" at 635,123 size 46x25; Text 'X'
   TextField "Campo de texto_53" at 633,181 size 46x25; Text 'Y'
   TextField "Campo de texto_54" at 636,239 size 46x25; Text 'Z'
   TextField "Campo de texto_55" at 506,79 size 284x25; Text 'MOMENTUKO X Y Z POSIZIOA'
   TextField "Campo de texto_56" at 14,304 size 448x25; Text 'MOMENTUKO ARDATZEN POSIZIOA GRADUTAN'
   Button "Botón_21" at 888,150 size 298x100; TextOff 'Pick & Place MARTXA'
      on Press: function_b14e0dd5("HMI_start", 0)
   Switch "Interruptor_1" at 52,70 size 64x32; CaptionText 'Switch'; TextOff 'OFF'; TextOn 'ON'
      on SwitchOn: SetBit("Power_DB_Power_a1")
      on SwitchOff: ResetBit("Power_DB_Power_a1")
   TextField "Campo de texto_57" at 52,45 size 87x25; Text 'Power A1'
   Switch "Interruptor_2" at 187,70 size 64x32; TextOn 'ON'; CaptionText 'Switch'; TextOff 'OFF'
      on SwitchOn: SetBit("Power_DB_Power_a2")
      on SwitchOff: ResetBit("Power_DB_Power_a2")
   TextField "Campo de texto_58" at 187,45 size 87x25; Text 'Power A2'
   Switch "Interruptor_3" at 322,70 size 64x32; TextOn 'ON'; CaptionText 'Switch'; TextOff 'OFF'
      on SwitchOff: ResetBit("Power_DB_Power_a3")
      on SwitchOn: SetBit("Power_DB_Power_a3")
   TextField "Campo de texto_59" at 322,45 size 87x25; Text 'Power A3'
   Switch "Interruptor_4" at 322,159 size 64x32; TextOn 'ON'; CaptionText 'Switch'; TextOff 'OFF'
      on SwitchOff: ResetBit("Tag_2")
      on SwitchOn: SetBit("Tag_2")
   Switch "Interruptor_5" at 322,207 size 64x32; TextOn 'ON'; CaptionText 'Switch'; TextOff 'OFF'
      on SwitchOff: ResetBit("Tag_3")
      on SwitchOn: SetBit("Tag_3")
   Switch "Interruptor_6" at 322,256 size 64x32; TextOn 'ON'; CaptionText 'Switch'; TextOff 'OFF'
      on SwitchOn: SetBit("Tag_6")
      on SwitchOff: ResetBit("Tag_6")
   TextField "Campo de texto_60" at 315,135 size 82x25; Text 'Freno A1'
   TextField "Campo de texto_61" at 315,187 size 82x25; Text 'Freno A2'
   TextField "Campo de texto_62" at 315,235 size 82x25; Text 'Freno A3'
   TextField "Campo de texto_33" at 952,334 size 241x25; Text 'MUGIMENDU ABSOLUTOAK'
   TextField "Campo de texto_40" at 569,568 size 290x23; Text 'Mugimendu absoluto point to point'
   Button "Botón_7" at 51,598 size 96x32; TextOff 'x+'
      on Press: function_b14e0dd5("x+", 0)
   Button "Botón_8" at 193,598 size 96x32; TextOff 'x-'
      on Press: function_b14e0dd5("x-", 0)
   Button "Botón_9" at 51,652 size 96x32; TextOff 'y+'
      on Press: function_b14e0dd5("y+", 0)
   Button "Botón_12" at 193,652 size 96x32; TextOff 'y-'
      on Press: function_b14e0dd5("y-", 0)
   Button "Botón_13" at 51,706 size 96x32; TextOff 'z+'
      on Press: function_b14e0dd5("z+", 0)
   Button "Botón_14" at 193,706 size 96x32; TextOff 'z-'
      on Press: function_b14e0dd5("z-", 0)
   Switch "Interruptor_7" at 132,529 size 64x32; CaptionText 'Switch'; TextOff 'OFF'; TextOn 'ON'
      on SwitchOn: SetBit("HABILITAR")
      on SwitchOff: ResetBit("HABILITAR")
   TextField "Campo de texto_34" at 116,490 size 100x25; Text 'JOG DELTA'
*)